(* Logix 5000 project; controller MV vendor 1 type 14 code 217 rev 31.11; software revision 31.00; part 27 of 53 *)
(* tags used below, declared in another part *)
   CWD : CHECKWORD_FLAGS;
   Dummy : BOOL;
   FVHR12_1701 : PlantItem;   // Valve FVHR12_17/01
   FVHR12_1702 : PlantItem;   // Valve FVHR12_17/02
   FVHR12_1703 : PlantItem;   // Valve FVHR12_17/03
   FVHR12_17_Valves_ON : BOOL;   // Check bit to confirm valves for FV12-17 route are open
   FVHR18_21_Valves_ON : BOOL;   // Check bit to confirm valves for FV18-21 route are open
   FVHR18_2501 : PlantItem;   // Valve FVHR18_25/01
   FVHR18_2502 : PlantItem;   // Valve FVHR18_25/02
   FVHR18_2503 : PlantItem;   // Valve FVHR18_25/03
   FVHR18_2504 : PlantItem;   // Valve FVHR18_25/04
   FVHR1_1101 : PlantItem;   // Valve FVHR1_11/01
   FVHR1_1102 : PlantItem;   // Valve FVHR1_11/02
   FVHR1_1103 : PlantItem;   // Valve FVHR1_11/03
   FVHR1_11_Valves_ON : BOOL;   // Check bit to confirm valves for FV1-11 route are open
   FVHR1_1701 : PlantItem;   // Valve FVHR1_17/01
   FVHR22_25_Valves_ON : BOOL;   // Check bit to confirm valves for FV22-25 route are open
   IGI_TestBit : BOOL;
   MC_B12 : INT[255];   // PX SWITCH Proxy switch flags f ile
   MC_B240 : INT[255];   // CH1 RN PMP Channel 1 return pum p drive flags
   MC_B241 : INT[255];   // CH2 RN PMP Channel 2 return pum p drive flags
   MC_B242 : INT[255];   // CH1 ROUTE Channel 1 route requ est flags
   MC_B243 : INT[255];   // CH2 ROUTE Channel 2 route requ est flags
   MC_B3 : INT[255];   // BINARY
   MC_bit_data_file_address : DINT;
   MC_bit_file_bit_offset : DINT;
   MC_bit_file_word_offset : DINT;
   MC_bit_offset : DINT;
   MC_bit_value_to_set : DINT;
   MC_CH2_CIP_BYPASS_Conditions : BOOL;
   MC_CH2_CIP_BYPASS_DrainConditions : BOOL;
   MC_CIP_AV01 : PlantItem;   // CIP_AV01
   MC_CIP_AV02 : PlantItem;   // CIP_AV02
   MC_CIP_AV05 : PlantItem;   // CIP_AV05
   MC_CIP_AV06 : PlantItem;   // CIP_AV06
   MC_CIP_AV07 : PlantItem;   // CIP_AV07
   MC_CIP_AV08 : PlantItem;   // CIP_AV08
   MC_CIP_AV09 : PlantItem;   // CIP_AV09
   MC_CIP_AV10 : PlantItem;   // CIP_AV10
   MC_CP1 : PlantItem;   // CP1
   MC_data_file_address : DINT;
   MC_GBYV1 : PlantItem;   // GBYV1
   MC_N10 : INT[255];   // SETTINGS
   MC_N100 : INT[255];   // C1_PLC Channel 1 PLC data
   MC_N101 : INT[255];   // CH1 PC>PLC Channel 1 PC to PLC
   MC_N102 : INT[255];   // CH1 PROG Channel 1 CIP progra m
   MC_N103 : INT[255];   // CH1 ITEMS Chwd.nos.of items to be checked for Chan nel 1
   MC_N104 : INT[255];   // CH1 REPORT Channel 1 CIP report file
   MC_N108 : INT[255];   // CH1 VDATA Channel 1 CIP progra m validation data
   MC_N112 : INT[255];   // FVR DATA Data read from FV ro uting PLC
   MC_N113 : INT[255];   // MVR DATA Data read from MV ro uting PLC
   MC_N114 : INT[255];   // YP DATA
   MC_N120 : INT[255];   // C2 PLC Channel 2 PLC data
   MC_N121 : INT[255];   // CH2 PC>PLC Channel 2 PC to PLC
   MC_N122 : INT[255];   // CH2 PROG Channel 2 CIP progra m
   MC_N123 : INT[255];   // CH2 ITEMS Chwd.nos.of items to be checked for Chan nel 2
   MC_N124 : INT[255];   // CH2 REPORT Channel 2 CIP report file
   MC_N128 : INT[255];   // CH2 VDATA Channel 2 CIP progra m validation data
   MC_N160 : INT[255];   // P40 CHECK
   MC_N161 : INT[255];   // P41 CHECK
   MC_N162 : INT[255];   // P42 CHECK
   MC_N163 : INT[255];   // P43 CHECK
   MC_N164 : INT[255];   // P44 CHECK
   MC_N165 : INT[255];   // P45 CHECK
   MC_N166 : INT[255];   // P46 CHECK
   MC_N167 : INT[255];   // Original N File From SLC, No Description Available
   MC_N20 : INT[255];   // P1 PRESS Control block and da ta for P1 pressure P ID loop
   MC_N200 : INT[255];   // CHK_WORK Plant item fault che cking work area
   MC_N201 : INT[255];   // P1 CHECK CIP program 1 plant item check list
   MC_N202 : INT[255];   // P2 CHECK CIP program 2 plant item check list
   MC_N203 : INT[255];   // P3 CHECK CIP program 3 plant item check list
   MC_N204 : INT[255];   // P4 CHECK CIP program 4 plant item check list
   MC_N205 : INT[255];   // P5 CHECK CIP program 5 plant item check list
   MC_N206 : INT[255];   // P6 CHECK CIP program 6 plant item check list
   MC_N207 : INT[255];   // P7 CHECK CIP program 7 plant item check list
   MC_N208 : INT[255];   // P8 CHECK CIP program 8 plant item check list
   MC_N209 : INT[255];   // P9 CHECK CIP program 9 plant item check list
   MC_N21 : INT[255];   // P1 FLOW Control block and da ta for P1 flowrate P ID loop
   MC_N210 : INT[255];   // P10 CHECK CIP program 10 plant item check list
   MC_N211 : INT[255];   // P11 CHECK CIP program 11 plant item check list
   MC_N212 : INT[255];   // P12 CHECK CIP program 12 plant item check list
   MC_N213 : INT[255];   // P13 CHECK CIP program 13 plant item check list
   MC_N214 : INT[255];   // P14 CHECK CIP program 14 plant item check list
   MC_N215 : INT[255];   // P15 CHECK CIP program 15 plant item check list
   MC_N216 : INT[255];   // P16 CHECK CIP program 16 plant item check list
   MC_N217 : INT[255];   // P17 CHECK CIP program 17 plant item check list
   MC_N218 : INT[255];   // P18 CHECK CIP program 18 plant item check list
   MC_N219 : INT[255];   // P19 CHECK CIP program 19 plant item check list
   MC_N22 : INT[255];   // P2 PRESS Control block and da ta for P2 pressure P ID loop
   MC_N220 : INT[255];   // P20 CHECK CIP program 20 plant item check list
   MC_N221 : INT[255];   // P21 CHECK CIP program 21 plant item check list
   MC_N222 : INT[255];   // P22 CHECK CIP program 22 plant item check list
   MC_N223 : INT[255];   // P23 CHECK CIP program 23 plant item check list
   MC_N224 : INT[255];   // P24 CHECK CIP program 24 plant item check list
   MC_N225 : INT[255];   // P25 CHECK CIP program 25 plant item check list
   MC_N226 : INT[255];   // P26 CHECK CIP program 26 plant item check list
   MC_N227 : INT[255];   // P27 CHECK CIP program 27 plant item check list
   MC_N228 : INT[255];   // P28 CHECK CIP program 28 plant item check list
   MC_N229 : INT[255];   // P29 CHECK CIP program 29 plant item check list
   MC_N23 : INT[255];   // P2 FLOW Control block and da ta for P2 flowrate P ID loop
   MC_N230 : INT[255];   // P30 CHECK CIP program 30 plant item check list
   MC_N231 : INT[255];   // P31 CHECK CIP program 31 plant item check list
   MC_N232 : INT[255];   // P32 CHECK CIP program 32 plant item check list
   MC_N233 : INT[255];   // P33 CHECK CIP program 33 plant item check list
   MC_N234 : INT[255];   // P34 CHECK CIP program 34 plant item check list
   MC_N235 : INT[255];   // P35 CHECK CIP program 35 plant item check list
   MC_N236 : INT[255];   // P36 CHECK CIP program 36 plant item check list
   MC_N237 : INT[255];   // P37 CHECK CIP program 37 plant item check list
   MC_N238 : INT[255];   // P38 CHECK CIP program 38 plant item check list
   MC_N239 : INT[255];   // P39 CHECK CIP program 39 plant item check list
   MC_N245 : INT[255];   // CC_WORK Continuous checking program work area
   MC_N255 : INT[255];   // CHECKWORDS Plant item checkword s
   MC_N7 : INT[255];   // INTEGER
   MC_N80 : INT[255];   // SRV1_PLC Detergent tank 1 ser vice PLC data
   MC_N81 : INT[255];   // SV1_PC Detergent tank 1 ser vice PC to PLC data
   MC_N82 : INT[255];   // SV1 ITEMS Chwd.nos.of items to be checked for DT1 service
   MC_N90 : INT[255];   // SV2_PLC Detergent tank 2 ser vice PLC data
   MC_N91 : INT[255];   // SV2_PC Detergent tank 2 ser vice PC to PLC data
   MC_N92 : INT[255];   // SV2 ITEMS Chwd.nos.of items to be checked for DT2 service
   MC_R3V1 : PlantItem;   // R3V1
   MC_SP_R1_1 : PlantItem;   // SP_R1_1
   MC_SP_R2_1 : PlantItem;   // SP_R2_1
   MC_SP_R2_2 : PlantItem;   // SP_R2_2
   MC_SP_R3_1 : PlantItem;   // SP_R3_1
   MC_SP_R5_1 : PlantItem;   // SP_R5_1
   MC_SP_R5_2 : PlantItem;   // SP_R5_2
   MC_SP_R6_1 : PlantItem;   // SP_R6_1
   MC_SP_R6_2 : PlantItem;   // SP_R6_2
   MC_SP_R6_3 : PlantItem;   // SP_R6_3
   MC_SP_R6_4 : PlantItem;   // SP_R6_4
   MC_SP_R6_5 : PlantItem;   // SP_R6_5
   MC_SP_V12TO17 : PlantItem;   // SP_V12TO17
   MC_SPV1 : PlantItem;   // SPV1
   MC_SPV2 : PlantItem;   // SPV2
   MC_SPV3 : PlantItem;   // SPV3
   MC_SPV4 : PlantItem;   // SPV4
   MC_SPV5 : PlantItem;   // SPV5
   MC_value_to_set : DINT;
   MC_word_offset : DINT;
(* MC_Common, continued *)

ROUTINE MC_Set_NFile_Value   (* ladder *)
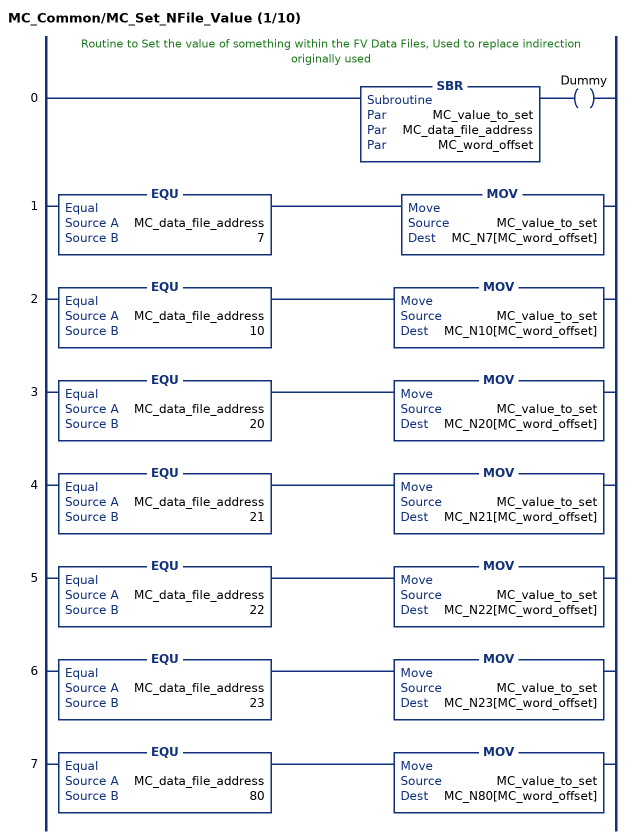
   // Routine to Set the value of something within the FV Data Files, Used to replace indirection originally used
   0: SBR(MC_value_to_set,MC_data_file_address,MC_word_offset)OTE(Dummy);
   1: EQU(MC_data_file_address,7)MOV(MC_value_to_set,MC_N7[MC_word_offset]);
   2: EQU(MC_data_file_address,10)MOV(MC_value_to_set,MC_N10[MC_word_offset]);
   3: EQU(MC_data_file_address,20)MOV(MC_value_to_set,MC_N20[MC_word_offset]);
   4: EQU(MC_data_file_address,21)MOV(MC_value_to_set,MC_N21[MC_word_offset]);
   5: EQU(MC_data_file_address,22)MOV(MC_value_to_set,MC_N22[MC_word_offset]);
   6: EQU(MC_data_file_address,23)MOV(MC_value_to_set,MC_N23[MC_word_offset]);
   7: EQU(MC_data_file_address,80)MOV(MC_value_to_set,MC_N80[MC_word_offset]);
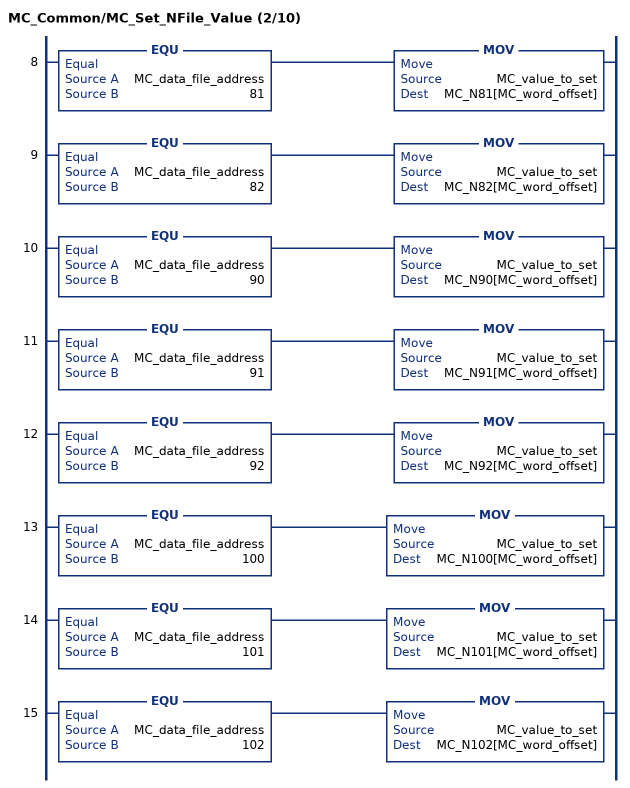
   8: EQU(MC_data_file_address,81)MOV(MC_value_to_set,MC_N81[MC_word_offset]);
   9: EQU(MC_data_file_address,82)MOV(MC_value_to_set,MC_N82[MC_word_offset]);
   10: EQU(MC_data_file_address,90)MOV(MC_value_to_set,MC_N90[MC_word_offset]);
   11: EQU(MC_data_file_address,91)MOV(MC_value_to_set,MC_N91[MC_word_offset]);
   12: EQU(MC_data_file_address,92)MOV(MC_value_to_set,MC_N92[MC_word_offset]);
   13: EQU(MC_data_file_address,100)MOV(MC_value_to_set,MC_N100[MC_word_offset]);
   14: EQU(MC_data_file_address,101)MOV(MC_value_to_set,MC_N101[MC_word_offset]);
   15: EQU(MC_data_file_address,102)MOV(MC_value_to_set,MC_N102[MC_word_offset]);
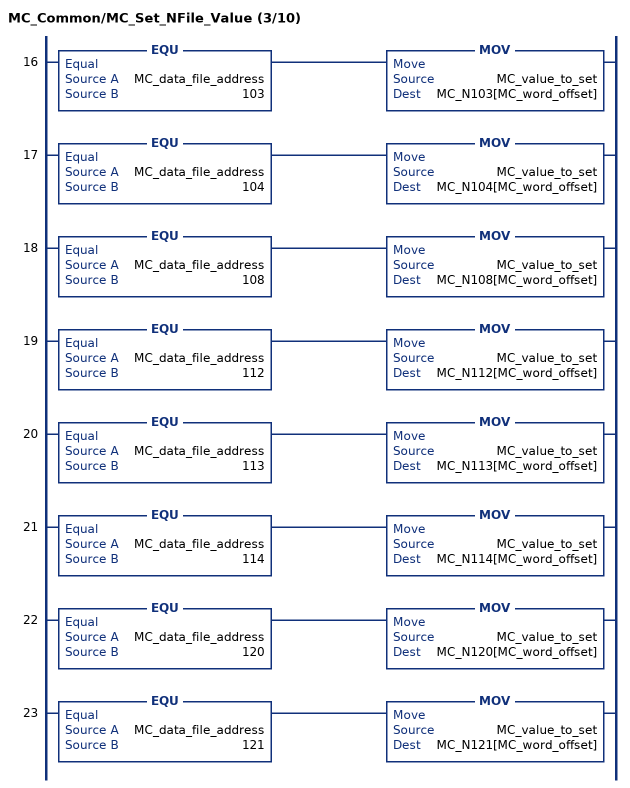
   16: EQU(MC_data_file_address,103)MOV(MC_value_to_set,MC_N103[MC_word_offset]);
   17: EQU(MC_data_file_address,104)MOV(MC_value_to_set,MC_N104[MC_word_offset]);
   18: EQU(MC_data_file_address,108)MOV(MC_value_to_set,MC_N108[MC_word_offset]);
   19: EQU(MC_data_file_address,112)MOV(MC_value_to_set,MC_N112[MC_word_offset]);
   20: EQU(MC_data_file_address,113)MOV(MC_value_to_set,MC_N113[MC_word_offset]);
   21: EQU(MC_data_file_address,114)MOV(MC_value_to_set,MC_N114[MC_word_offset]);
   22: EQU(MC_data_file_address,120)MOV(MC_value_to_set,MC_N120[MC_word_offset]);
   23: EQU(MC_data_file_address,121)MOV(MC_value_to_set,MC_N121[MC_word_offset]);
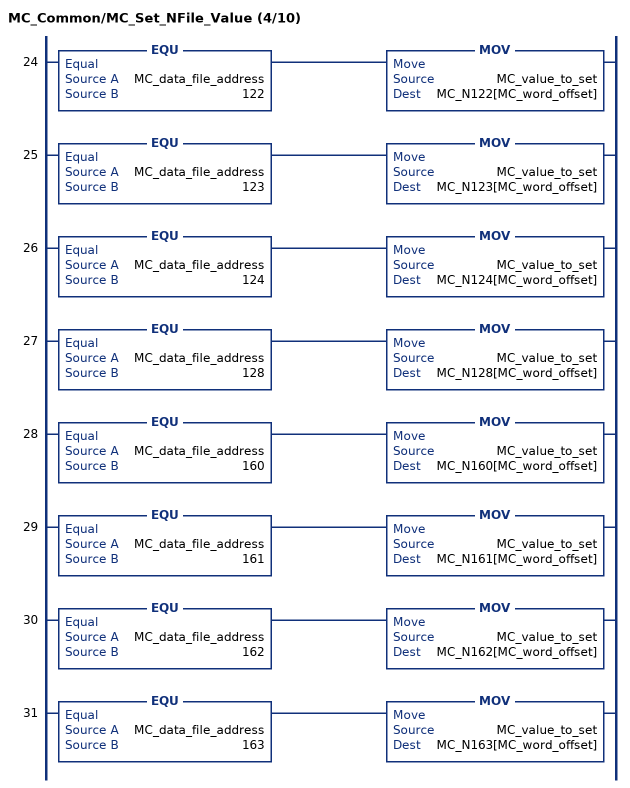
   24: EQU(MC_data_file_address,122)MOV(MC_value_to_set,MC_N122[MC_word_offset]);
   25: EQU(MC_data_file_address,123)MOV(MC_value_to_set,MC_N123[MC_word_offset]);
   26: EQU(MC_data_file_address,124)MOV(MC_value_to_set,MC_N124[MC_word_offset]);
   27: EQU(MC_data_file_address,128)MOV(MC_value_to_set,MC_N128[MC_word_offset]);
   28: EQU(MC_data_file_address,160)MOV(MC_value_to_set,MC_N160[MC_word_offset]);
   29: EQU(MC_data_file_address,161)MOV(MC_value_to_set,MC_N161[MC_word_offset]);
   30: EQU(MC_data_file_address,162)MOV(MC_value_to_set,MC_N162[MC_word_offset]);
   31: EQU(MC_data_file_address,163)MOV(MC_value_to_set,MC_N163[MC_word_offset]);
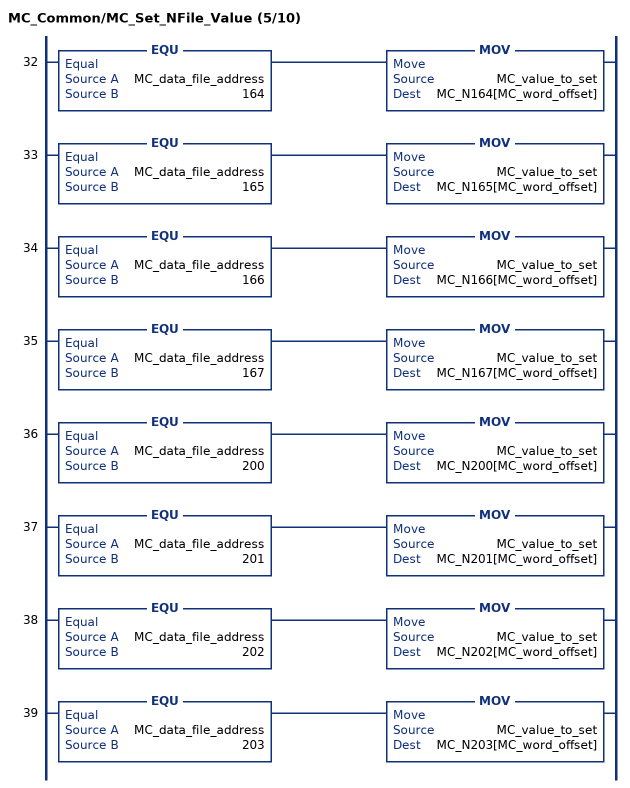
   32: EQU(MC_data_file_address,164)MOV(MC_value_to_set,MC_N164[MC_word_offset]);
   33: EQU(MC_data_file_address,165)MOV(MC_value_to_set,MC_N165[MC_word_offset]);
   34: EQU(MC_data_file_address,166)MOV(MC_value_to_set,MC_N166[MC_word_offset]);
   35: EQU(MC_data_file_address,167)MOV(MC_value_to_set,MC_N167[MC_word_offset]);
   36: EQU(MC_data_file_address,200)MOV(MC_value_to_set,MC_N200[MC_word_offset]);
   37: EQU(MC_data_file_address,201)MOV(MC_value_to_set,MC_N201[MC_word_offset]);
   38: EQU(MC_data_file_address,202)MOV(MC_value_to_set,MC_N202[MC_word_offset]);
   39: EQU(MC_data_file_address,203)MOV(MC_value_to_set,MC_N203[MC_word_offset]);
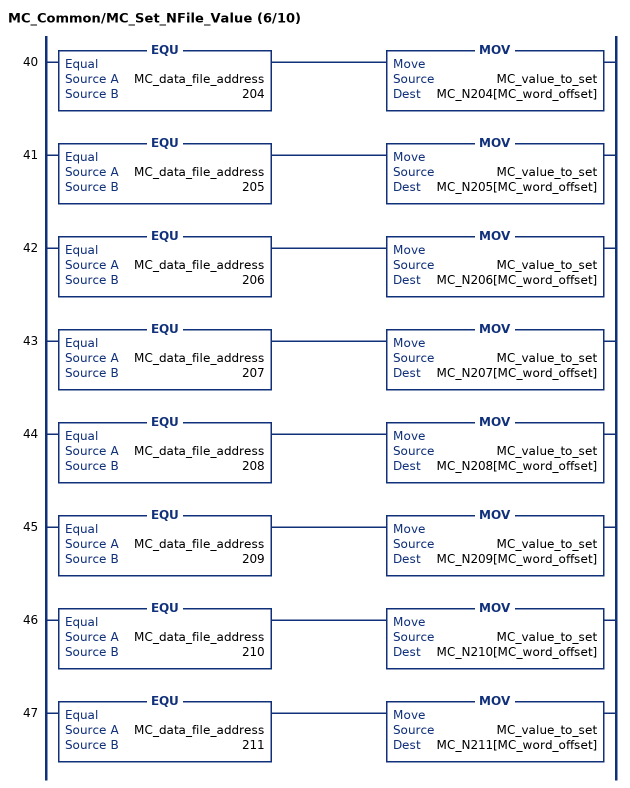
   40: EQU(MC_data_file_address,204)MOV(MC_value_to_set,MC_N204[MC_word_offset]);
   41: EQU(MC_data_file_address,205)MOV(MC_value_to_set,MC_N205[MC_word_offset]);
   42: EQU(MC_data_file_address,206)MOV(MC_value_to_set,MC_N206[MC_word_offset]);
   43: EQU(MC_data_file_address,207)MOV(MC_value_to_set,MC_N207[MC_word_offset]);
   44: EQU(MC_data_file_address,208)MOV(MC_value_to_set,MC_N208[MC_word_offset]);
   45: EQU(MC_data_file_address,209)MOV(MC_value_to_set,MC_N209[MC_word_offset]);
   46: EQU(MC_data_file_address,210)MOV(MC_value_to_set,MC_N210[MC_word_offset]);
   47: EQU(MC_data_file_address,211)MOV(MC_value_to_set,MC_N211[MC_word_offset]);
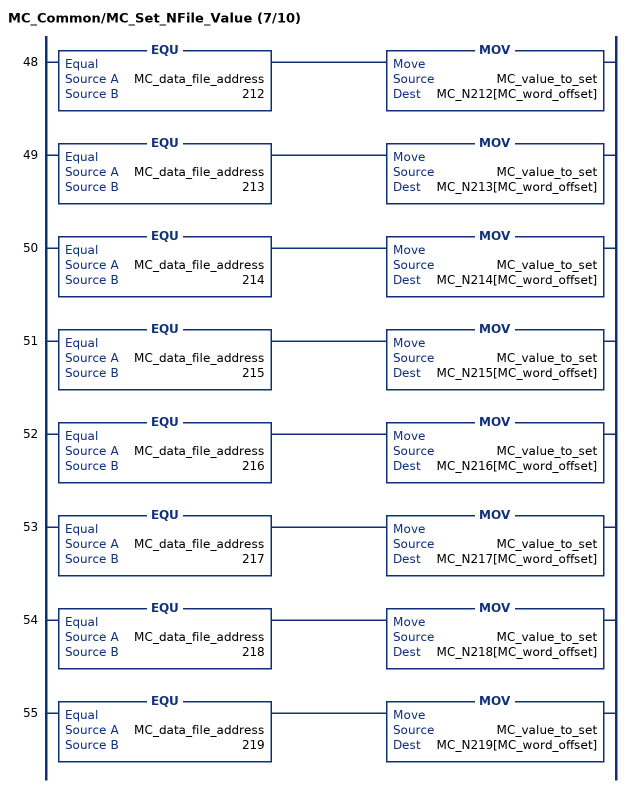
   48: EQU(MC_data_file_address,212)MOV(MC_value_to_set,MC_N212[MC_word_offset]);
   49: EQU(MC_data_file_address,213)MOV(MC_value_to_set,MC_N213[MC_word_offset]);
   50: EQU(MC_data_file_address,214)MOV(MC_value_to_set,MC_N214[MC_word_offset]);
   51: EQU(MC_data_file_address,215)MOV(MC_value_to_set,MC_N215[MC_word_offset]);
   52: EQU(MC_data_file_address,216)MOV(MC_value_to_set,MC_N216[MC_word_offset]);
   53: EQU(MC_data_file_address,217)MOV(MC_value_to_set,MC_N217[MC_word_offset]);
   54: EQU(MC_data_file_address,218)MOV(MC_value_to_set,MC_N218[MC_word_offset]);
   55: EQU(MC_data_file_address,219)MOV(MC_value_to_set,MC_N219[MC_word_offset]);
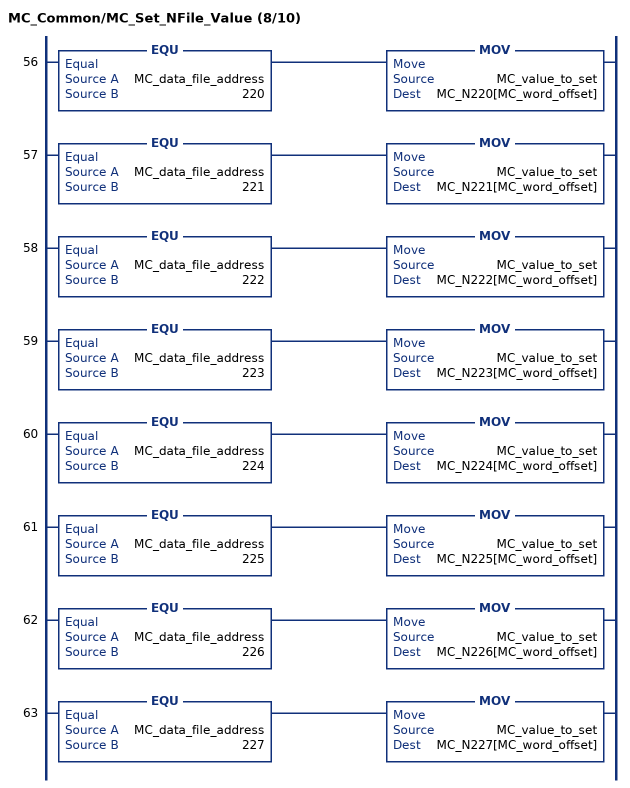
   56: EQU(MC_data_file_address,220)MOV(MC_value_to_set,MC_N220[MC_word_offset]);
   57: EQU(MC_data_file_address,221)MOV(MC_value_to_set,MC_N221[MC_word_offset]);
   58: EQU(MC_data_file_address,222)MOV(MC_value_to_set,MC_N222[MC_word_offset]);
   59: EQU(MC_data_file_address,223)MOV(MC_value_to_set,MC_N223[MC_word_offset]);
   60: EQU(MC_data_file_address,224)MOV(MC_value_to_set,MC_N224[MC_word_offset]);
   61: EQU(MC_data_file_address,225)MOV(MC_value_to_set,MC_N225[MC_word_offset]);
   62: EQU(MC_data_file_address,226)MOV(MC_value_to_set,MC_N226[MC_word_offset]);
   63: EQU(MC_data_file_address,227)MOV(MC_value_to_set,MC_N227[MC_word_offset]);
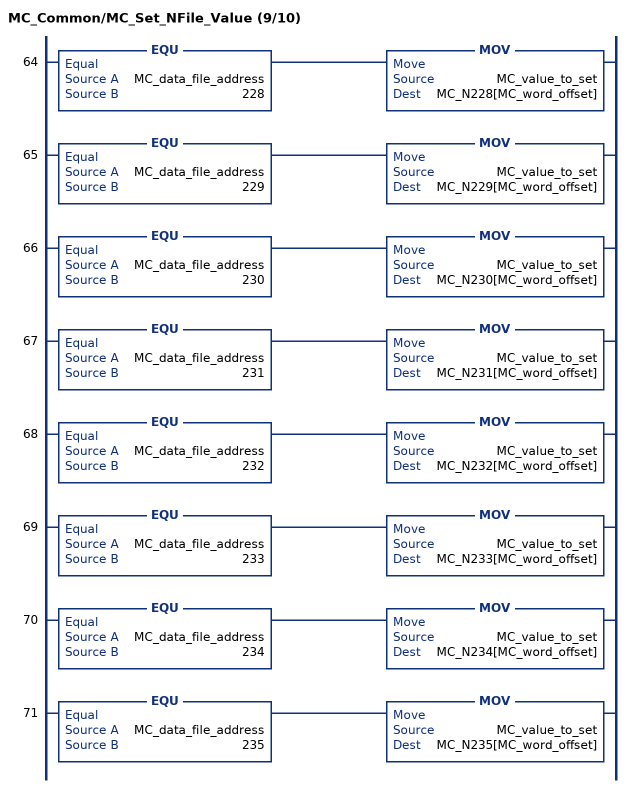
   64: EQU(MC_data_file_address,228)MOV(MC_value_to_set,MC_N228[MC_word_offset]);
   65: EQU(MC_data_file_address,229)MOV(MC_value_to_set,MC_N229[MC_word_offset]);
   66: EQU(MC_data_file_address,230)MOV(MC_value_to_set,MC_N230[MC_word_offset]);
   67: EQU(MC_data_file_address,231)MOV(MC_value_to_set,MC_N231[MC_word_offset]);
   68: EQU(MC_data_file_address,232)MOV(MC_value_to_set,MC_N232[MC_word_offset]);
   69: EQU(MC_data_file_address,233)MOV(MC_value_to_set,MC_N233[MC_word_offset]);
   70: EQU(MC_data_file_address,234)MOV(MC_value_to_set,MC_N234[MC_word_offset]);
   71: EQU(MC_data_file_address,235)MOV(MC_value_to_set,MC_N235[MC_word_offset]);
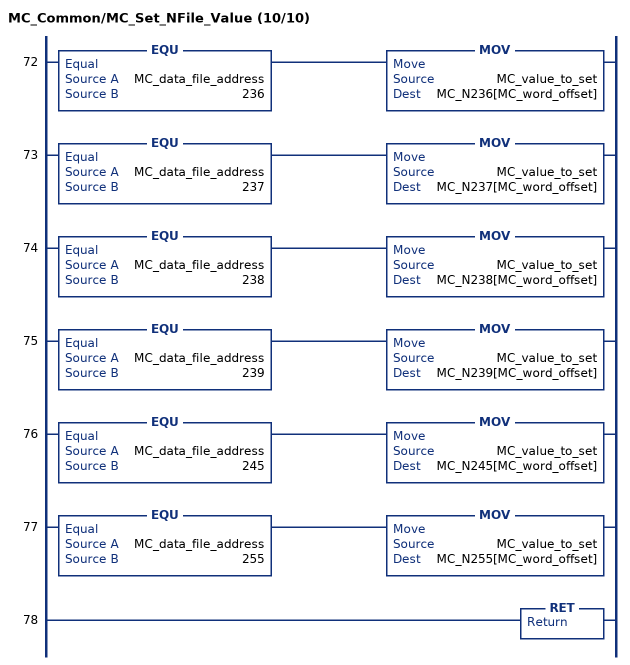
   72: EQU(MC_data_file_address,236)MOV(MC_value_to_set,MC_N236[MC_word_offset]);
   73: EQU(MC_data_file_address,237)MOV(MC_value_to_set,MC_N237[MC_word_offset]);
   74: EQU(MC_data_file_address,238)MOV(MC_value_to_set,MC_N238[MC_word_offset]);
   75: EQU(MC_data_file_address,239)MOV(MC_value_to_set,MC_N239[MC_word_offset]);
   76: EQU(MC_data_file_address,245)MOV(MC_value_to_set,MC_N245[MC_word_offset]);
   77: EQU(MC_data_file_address,255)MOV(MC_value_to_set,MC_N255[MC_word_offset]);
   78: RET();
END_ROUTINE

ROUTINE MC_SetBitFile_Value   (* ladder *)
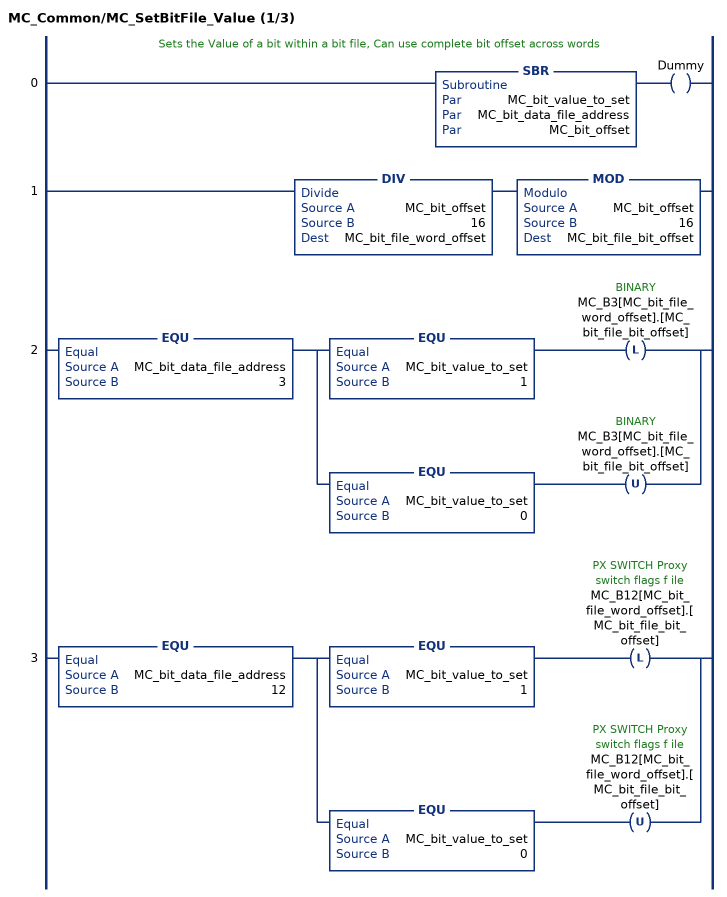
   // Sets the Value of a bit within a bit file, Can use complete bit offset across words
   0: SBR(MC_bit_value_to_set,MC_bit_data_file_address,MC_bit_offset)OTE(Dummy);
   1: DIV(MC_bit_offset,16,MC_bit_file_word_offset)MOD(MC_bit_offset,16,MC_bit_file_bit_offset);
   2: EQU(MC_bit_data_file_address,3)[EQU(MC_bit_value_to_set,1) OTL(MC_B3[MC_bit_file_word_offset].[MC_bit_file_bit_offset]) ,EQU(MC_bit_value_to_set,0) OTU(MC_B3[MC_bit_file_word_offset].[MC_bit_file_bit_offset]) ];
   3: EQU(MC_bit_data_file_address,12)[EQU(MC_bit_value_to_set,1) OTL(MC_B12[MC_bit_file_word_offset].[MC_bit_file_bit_offset]) ,EQU(MC_bit_value_to_set,0) OTU(MC_B12[MC_bit_file_word_offset].[MC_bit_file_bit_offset]) ];
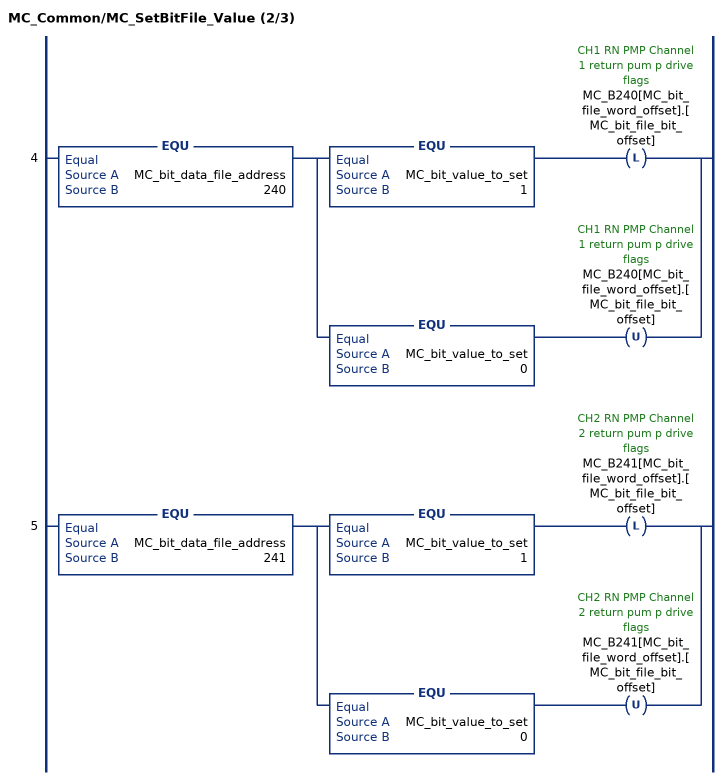
   4: EQU(MC_bit_data_file_address,240)[EQU(MC_bit_value_to_set,1) OTL(MC_B240[MC_bit_file_word_offset].[MC_bit_file_bit_offset]) ,EQU(MC_bit_value_to_set,0) OTU(MC_B240[MC_bit_file_word_offset].[MC_bit_file_bit_offset]) ];
   5: EQU(MC_bit_data_file_address,241)[EQU(MC_bit_value_to_set,1) OTL(MC_B241[MC_bit_file_word_offset].[MC_bit_file_bit_offset]) ,EQU(MC_bit_value_to_set,0) OTU(MC_B241[MC_bit_file_word_offset].[MC_bit_file_bit_offset]) ];
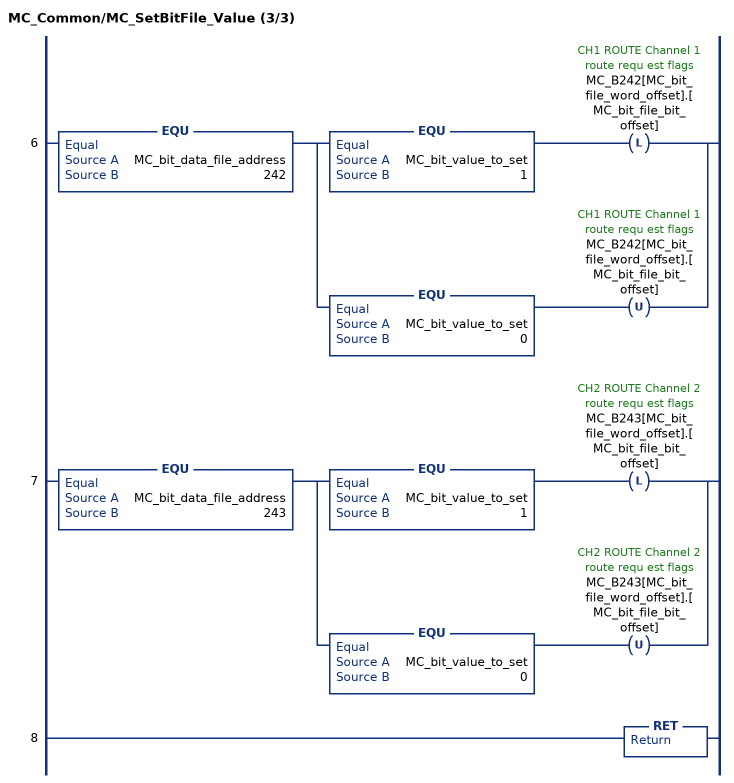
   6: EQU(MC_bit_data_file_address,242)[EQU(MC_bit_value_to_set,1) OTL(MC_B242[MC_bit_file_word_offset].[MC_bit_file_bit_offset]) ,EQU(MC_bit_value_to_set,0) OTU(MC_B242[MC_bit_file_word_offset].[MC_bit_file_bit_offset]) ];
   7: EQU(MC_bit_data_file_address,243)[EQU(MC_bit_value_to_set,1) OTL(MC_B243[MC_bit_file_word_offset].[MC_bit_file_bit_offset]) ,EQU(MC_bit_value_to_set,0) OTU(MC_B243[MC_bit_file_word_offset].[MC_bit_file_bit_offset]) ];
   8: RET();
END_ROUTINE

ROUTINE MC_SHARE_ITEM_240   (* ladder *)
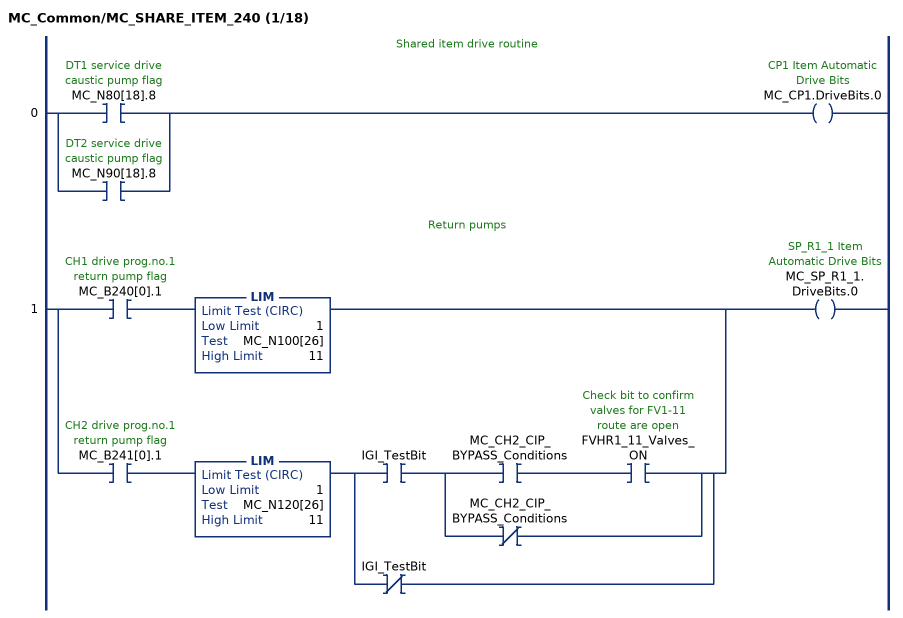
   // Shared item drive routine
   0: [XIC(MC_N80[18].8) ,XIC(MC_N90[18].8) ]OTE(MC_CP1.DriveBits.0);
   // Return pumps
   1: [XIC(MC_B240[0].1) LIM(1,MC_N100[26],11) ,XIC(MC_B241[0].1) LIM(1,MC_N120[26],11) [XIC(IGI_TestBit) [XIC(MC_CH2_CIP_BYPASS_Conditions) XIC(FVHR1_11_Valves_ON) ,XIO(MC_CH2_CIP_BYPASS_Conditions) ] ,XIO(IGI_TestBit) ] ]OTE(MC_SP_R1_1.DriveBits.0);
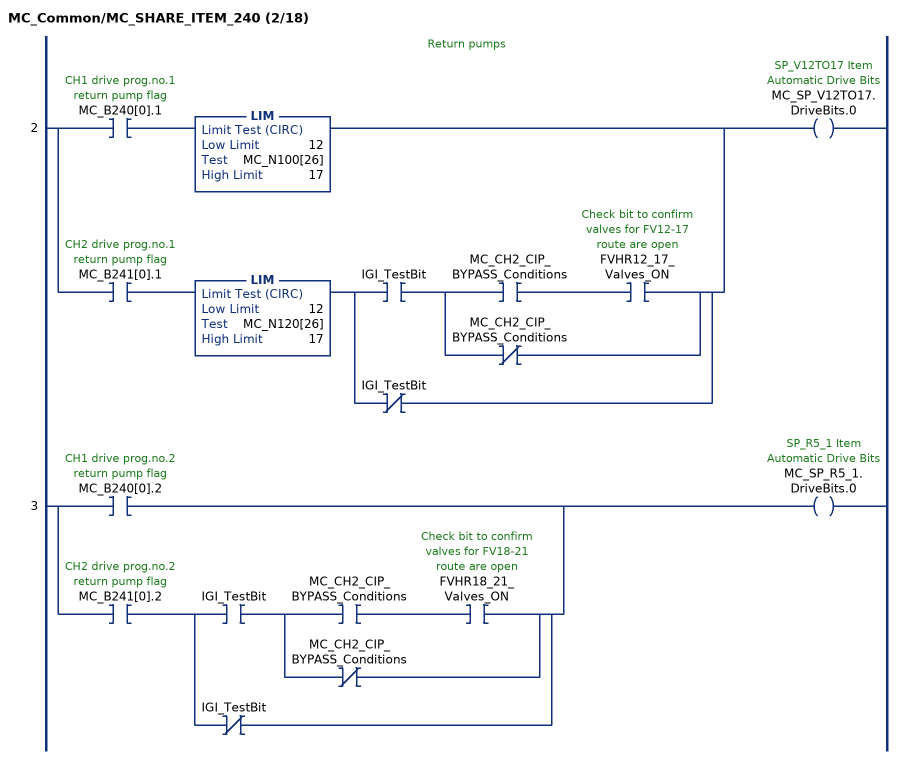
   // Return pumps
   2: [XIC(MC_B240[0].1) LIM(12,MC_N100[26],17) ,XIC(MC_B241[0].1) LIM(12,MC_N120[26],17) [XIC(IGI_TestBit) [XIC(MC_CH2_CIP_BYPASS_Conditions) XIC(FVHR12_17_Valves_ON) ,XIO(MC_CH2_CIP_BYPASS_Conditions) ] ,XIO(IGI_TestBit) ] ]OTE(MC_SP_V12TO17.DriveBits.0);
   3: [XIC(MC_B240[0].2) ,XIC(MC_B241[0].2) [XIC(IGI_TestBit) [XIC(MC_CH2_CIP_BYPASS_Conditions) XIC(FVHR18_21_Valves_ON) ,XIO(MC_CH2_CIP_BYPASS_Conditions) ] ,XIO(IGI_TestBit) ] ]OTE(MC_SP_R5_1.DriveBits.0);
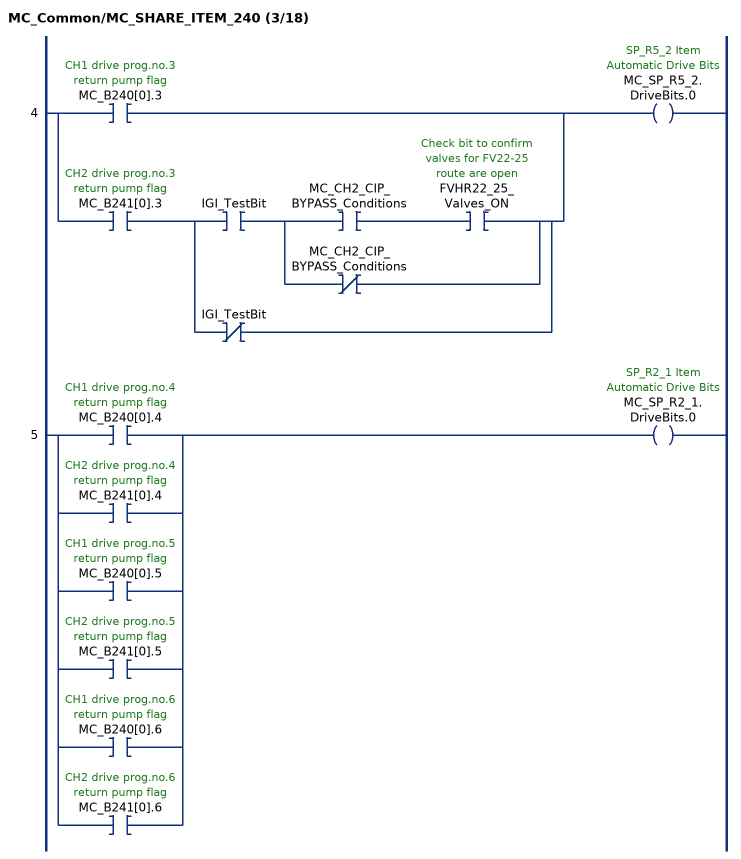
   4: [XIC(MC_B240[0].3) ,XIC(MC_B241[0].3) [XIC(IGI_TestBit) [XIC(MC_CH2_CIP_BYPASS_Conditions) XIC(FVHR22_25_Valves_ON) ,XIO(MC_CH2_CIP_BYPASS_Conditions) ] ,XIO(IGI_TestBit) ] ]OTE(MC_SP_R5_2.DriveBits.0);
   5: [XIC(MC_B240[0].4) ,XIC(MC_B241[0].4) ,XIC(MC_B240[0].5) ,XIC(MC_B241[0].5) ,XIC(MC_B240[0].6) ,XIC(MC_B241[0].6) ]OTE(MC_SP_R2_1.DriveBits.0);
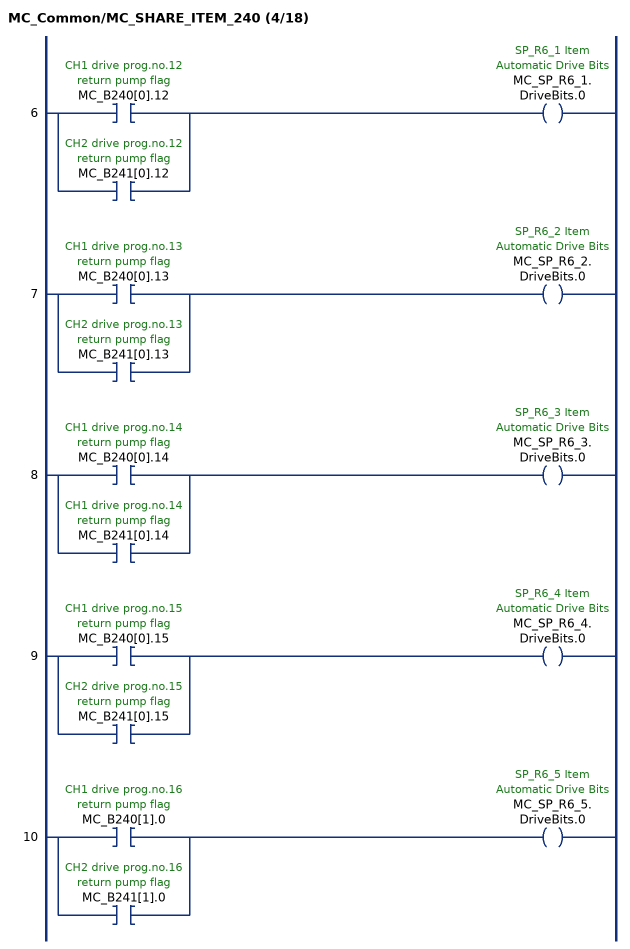
   6: [XIC(MC_B240[0].12) ,XIC(MC_B241[0].12) ]OTE(MC_SP_R6_1.DriveBits.0);
   7: [XIC(MC_B240[0].13) ,XIC(MC_B241[0].13) ]OTE(MC_SP_R6_2.DriveBits.0);
   8: [XIC(MC_B240[0].14) ,XIC(MC_B241[0].14) ]OTE(MC_SP_R6_3.DriveBits.0);
   9: [XIC(MC_B240[0].15) ,XIC(MC_B241[0].15) ]OTE(MC_SP_R6_4.DriveBits.0);
   10: [XIC(MC_B240[1].0) ,XIC(MC_B241[1].0) ]OTE(MC_SP_R6_5.DriveBits.0);
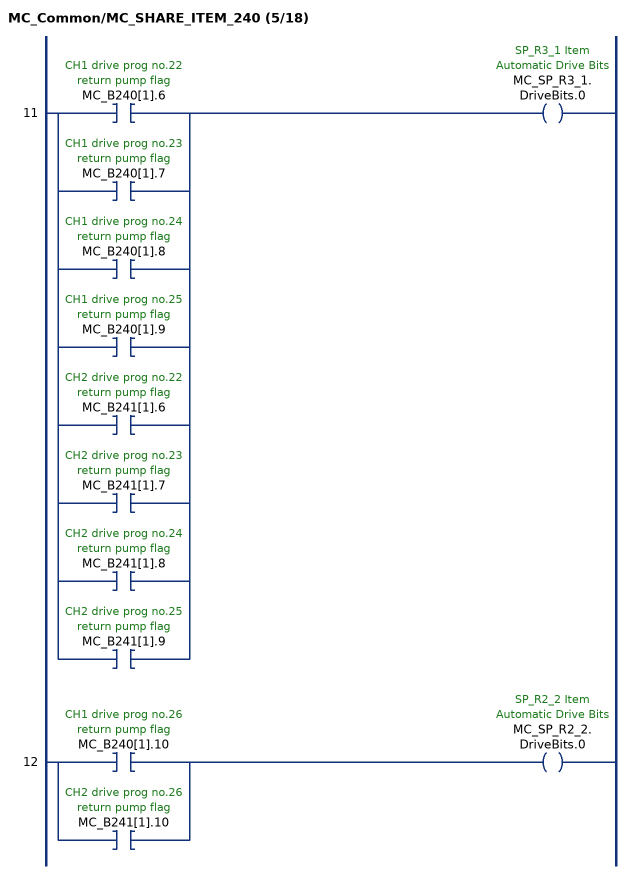
   11: [XIC(MC_B240[1].6) ,XIC(MC_B240[1].7) ,XIC(MC_B240[1].8) ,XIC(MC_B240[1].9) ,XIC(MC_B241[1].6) ,XIC(MC_B241[1].7) ,XIC(MC_B241[1].8) ,XIC(MC_B241[1].9) ]OTE(MC_SP_R3_1.DriveBits.0);
   12: [XIC(MC_B240[1].10) ,XIC(MC_B241[1].10) ]OTE(MC_SP_R2_2.DriveBits.0);
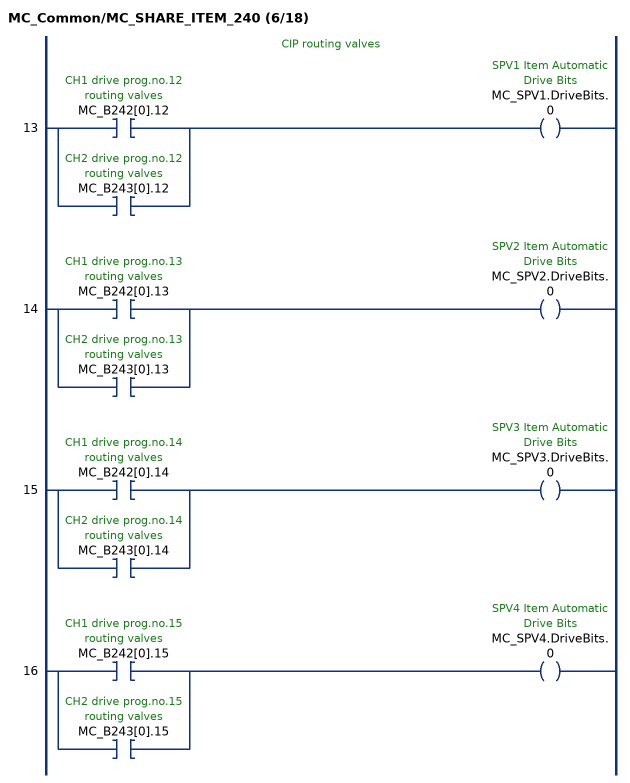
   // CIP routing valves
   13: [XIC(MC_B242[0].12) ,XIC(MC_B243[0].12) ]OTE(MC_SPV1.DriveBits.0);
   14: [XIC(MC_B242[0].13) ,XIC(MC_B243[0].13) ]OTE(MC_SPV2.DriveBits.0);
   15: [XIC(MC_B242[0].14) ,XIC(MC_B243[0].14) ]OTE(MC_SPV3.DriveBits.0);
   16: [XIC(MC_B242[0].15) ,XIC(MC_B243[0].15) ]OTE(MC_SPV4.DriveBits.0);
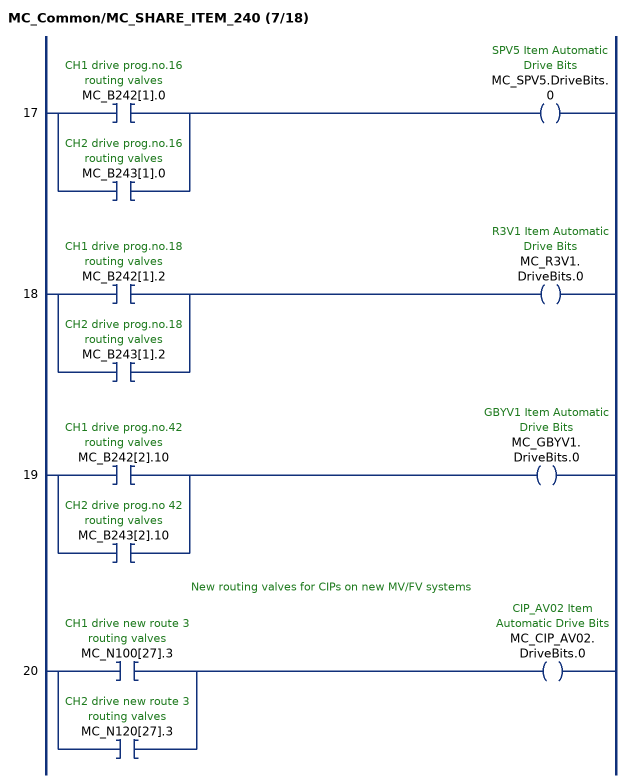
   17: [XIC(MC_B242[1].0) ,XIC(MC_B243[1].0) ]OTE(MC_SPV5.DriveBits.0);
   18: [XIC(MC_B242[1].2) ,XIC(MC_B243[1].2) ]OTE(MC_R3V1.DriveBits.0);
   19: [XIC(MC_B242[2].10) ,XIC(MC_B243[2].10) ]OTE(MC_GBYV1.DriveBits.0);
   // New routing valves for CIPs on new MV/FV systems
   20: [XIC(MC_N100[27].3) ,XIC(MC_N120[27].3) ]OTE(MC_CIP_AV02.DriveBits.0);
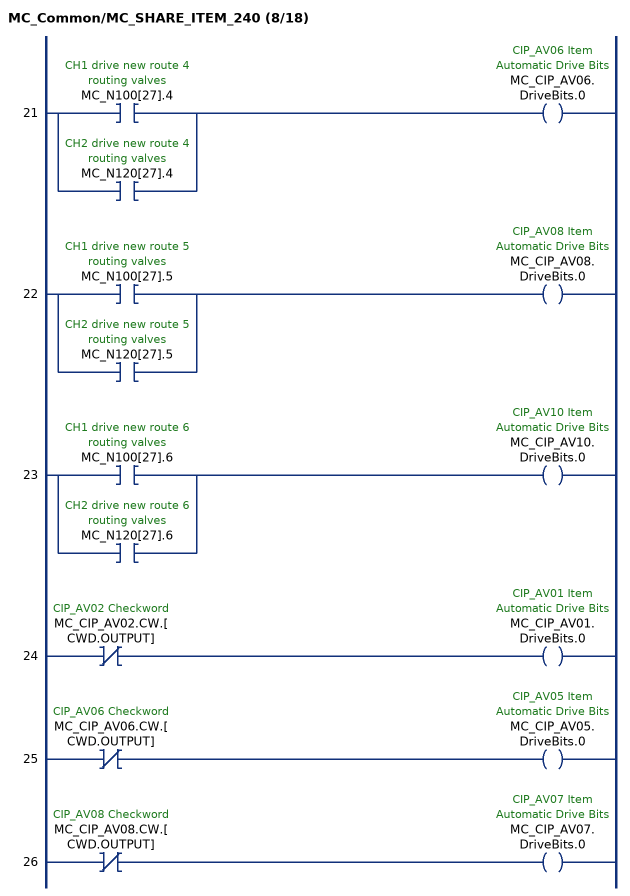
   21: [XIC(MC_N100[27].4) ,XIC(MC_N120[27].4) ]OTE(MC_CIP_AV06.DriveBits.0);
   22: [XIC(MC_N100[27].5) ,XIC(MC_N120[27].5) ]OTE(MC_CIP_AV08.DriveBits.0);
   23: [XIC(MC_N100[27].6) ,XIC(MC_N120[27].6) ]OTE(MC_CIP_AV10.DriveBits.0);
   24: XIO(MC_CIP_AV02.CW.[CWD.OUTPUT])OTE(MC_CIP_AV01.DriveBits.0);
   25: XIO(MC_CIP_AV06.CW.[CWD.OUTPUT])OTE(MC_CIP_AV05.DriveBits.0);
   26: XIO(MC_CIP_AV08.CW.[CWD.OUTPUT])OTE(MC_CIP_AV07.DriveBits.0);
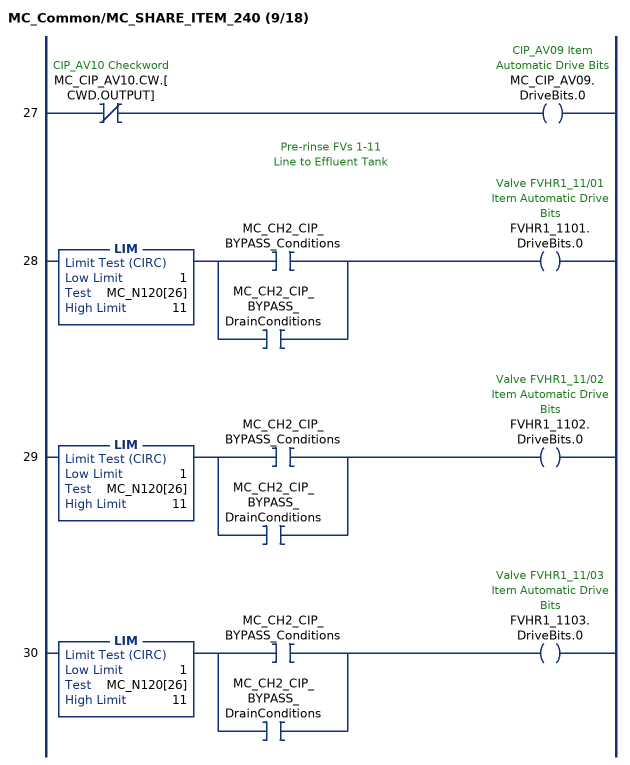
   27: XIO(MC_CIP_AV10.CW.[CWD.OUTPUT])OTE(MC_CIP_AV09.DriveBits.0);
   // Pre-rinse FVs 1-11
   // Line to Effluent Tank
   28: LIM(1,MC_N120[26],11)[XIC(MC_CH2_CIP_BYPASS_Conditions) ,XIC(MC_CH2_CIP_BYPASS_DrainConditions) ]OTE(FVHR1_1101.DriveBits.0);
   29: LIM(1,MC_N120[26],11)[XIC(MC_CH2_CIP_BYPASS_Conditions) ,XIC(MC_CH2_CIP_BYPASS_DrainConditions) ]OTE(FVHR1_1102.DriveBits.0);
   30: LIM(1,MC_N120[26],11)[XIC(MC_CH2_CIP_BYPASS_Conditions) ,XIC(MC_CH2_CIP_BYPASS_DrainConditions) ]OTE(FVHR1_1103.DriveBits.0);
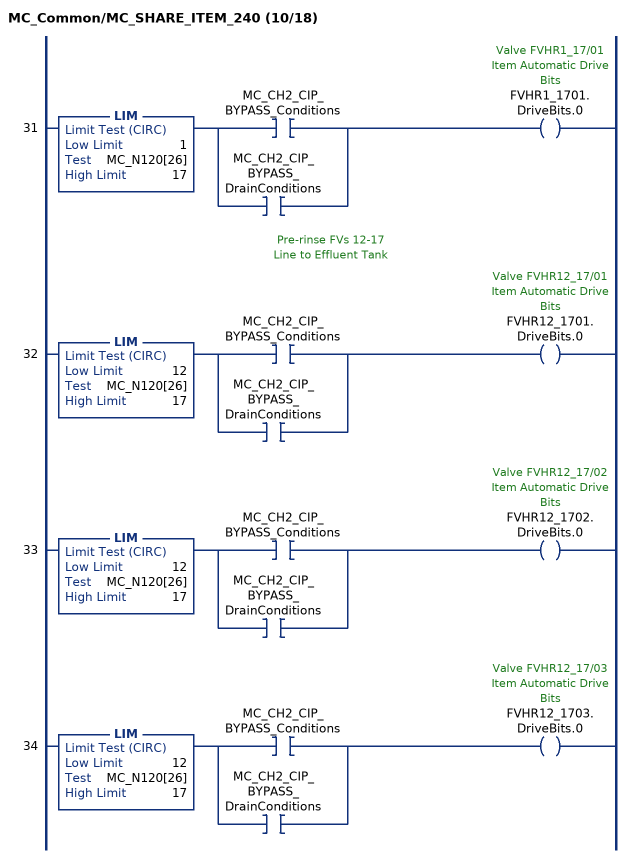
   31: LIM(1,MC_N120[26],17)[XIC(MC_CH2_CIP_BYPASS_Conditions) ,XIC(MC_CH2_CIP_BYPASS_DrainConditions) ]OTE(FVHR1_1701.DriveBits.0);
   // Pre-rinse FVs 12-17
   // Line to Effluent Tank
   32: LIM(12,MC_N120[26],17)[XIC(MC_CH2_CIP_BYPASS_Conditions) ,XIC(MC_CH2_CIP_BYPASS_DrainConditions) ]OTE(FVHR12_1701.DriveBits.0);
   33: LIM(12,MC_N120[26],17)[XIC(MC_CH2_CIP_BYPASS_Conditions) ,XIC(MC_CH2_CIP_BYPASS_DrainConditions) ]OTE(FVHR12_1702.DriveBits.0);
   34: LIM(12,MC_N120[26],17)[XIC(MC_CH2_CIP_BYPASS_Conditions) ,XIC(MC_CH2_CIP_BYPASS_DrainConditions) ]OTE(FVHR12_1703.DriveBits.0);
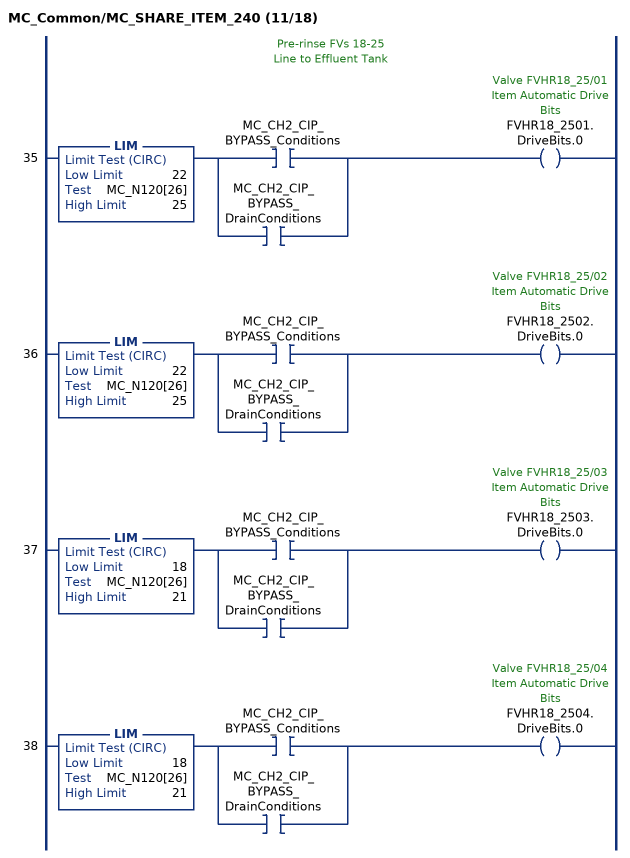
   // Pre-rinse FVs 18-25
   // Line to Effluent Tank
   35: LIM(22,MC_N120[26],25)[XIC(MC_CH2_CIP_BYPASS_Conditions) ,XIC(MC_CH2_CIP_BYPASS_DrainConditions) ]OTE(FVHR18_2501.DriveBits.0);
   36: LIM(22,MC_N120[26],25)[XIC(MC_CH2_CIP_BYPASS_Conditions) ,XIC(MC_CH2_CIP_BYPASS_DrainConditions) ]OTE(FVHR18_2502.DriveBits.0);
   37: LIM(18,MC_N120[26],21)[XIC(MC_CH2_CIP_BYPASS_Conditions) ,XIC(MC_CH2_CIP_BYPASS_DrainConditions) ]OTE(FVHR18_2503.DriveBits.0);
   38: LIM(18,MC_N120[26],21)[XIC(MC_CH2_CIP_BYPASS_Conditions) ,XIC(MC_CH2_CIP_BYPASS_DrainConditions) ]OTE(FVHR18_2504.DriveBits.0);
